REGION Network 277: SAFE OUTPUT CARD FAULT
   RUNG wire#powerrail
      Contact( "reset" )
      { S7_Templates := "SrcType := Word" } EQ_Contact(in1 := "DB101_DB_SDC_FAULTS".Carrier_Fault[28], in2 := 122)
      Coil( "DB302_HMI_Faults".Carrier28_Faults_0.%X9 )
   END_RUNG
   // the same network as SCL:
   "DB302_HMI_Faults".Carrier28_Faults_0.%X9 := "reset" AND ("DB101_DB_SDC_FAULTS".Carrier_Fault[28] = 122);
END_REGION

REGION Network 278: STANDARD INPUT CARD FAULT
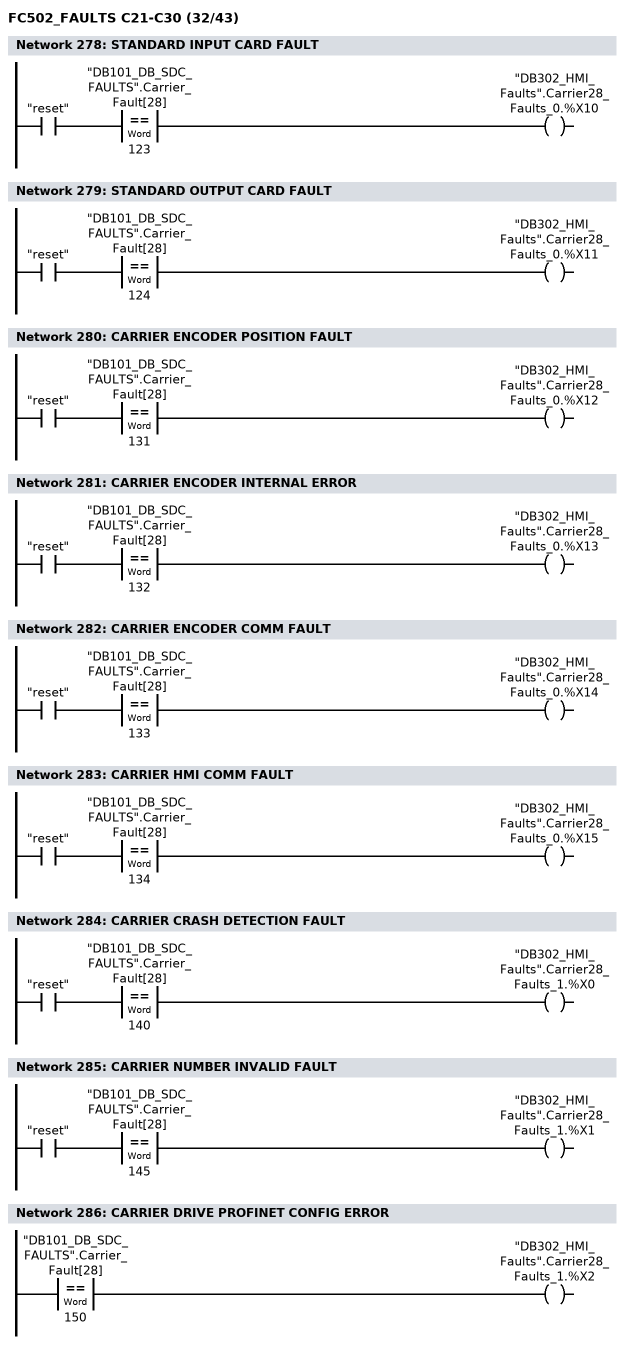
   RUNG wire#powerrail
      Contact( "reset" )
      { S7_Templates := "SrcType := Word" } EQ_Contact(in1 := "DB101_DB_SDC_FAULTS".Carrier_Fault[28], in2 := 123)
      Coil( "DB302_HMI_Faults".Carrier28_Faults_0.%X10 )
   END_RUNG
   // the same network as SCL:
   "DB302_HMI_Faults".Carrier28_Faults_0.%X10 := "reset" AND ("DB101_DB_SDC_FAULTS".Carrier_Fault[28] = 123);
END_REGION

REGION Network 279: STANDARD OUTPUT CARD FAULT
   RUNG wire#powerrail
      Contact( "reset" )
      { S7_Templates := "SrcType := Word" } EQ_Contact(in1 := "DB101_DB_SDC_FAULTS".Carrier_Fault[28], in2 := 124)
      Coil( "DB302_HMI_Faults".Carrier28_Faults_0.%X11 )
   END_RUNG
   // the same network as SCL:
   "DB302_HMI_Faults".Carrier28_Faults_0.%X11 := "reset" AND ("DB101_DB_SDC_FAULTS".Carrier_Fault[28] = 124);
END_REGION

REGION Network 280: CARRIER ENCODER POSITION FAULT
   RUNG wire#powerrail
      Contact( "reset" )
      { S7_Templates := "SrcType := Word" } EQ_Contact(in1 := "DB101_DB_SDC_FAULTS".Carrier_Fault[28], in2 := 131)
      Coil( "DB302_HMI_Faults".Carrier28_Faults_0.%X12 )
   END_RUNG
   // the same network as SCL:
   "DB302_HMI_Faults".Carrier28_Faults_0.%X12 := "reset" AND ("DB101_DB_SDC_FAULTS".Carrier_Fault[28] = 131);
END_REGION

REGION Network 281: CARRIER ENCODER INTERNAL ERROR
   RUNG wire#powerrail
      Contact( "reset" )
      { S7_Templates := "SrcType := Word" } EQ_Contact(in1 := "DB101_DB_SDC_FAULTS".Carrier_Fault[28], in2 := 132)
      Coil( "DB302_HMI_Faults".Carrier28_Faults_0.%X13 )
   END_RUNG
   // the same network as SCL:
   "DB302_HMI_Faults".Carrier28_Faults_0.%X13 := "reset" AND ("DB101_DB_SDC_FAULTS".Carrier_Fault[28] = 132);
END_REGION

REGION Network 282: CARRIER ENCODER COMM FAULT
   RUNG wire#powerrail
      Contact( "reset" )
      { S7_Templates := "SrcType := Word" } EQ_Contact(in1 := "DB101_DB_SDC_FAULTS".Carrier_Fault[28], in2 := 133)
      Coil( "DB302_HMI_Faults".Carrier28_Faults_0.%X14 )
   END_RUNG
   // the same network as SCL:
   "DB302_HMI_Faults".Carrier28_Faults_0.%X14 := "reset" AND ("DB101_DB_SDC_FAULTS".Carrier_Fault[28] = 133);
END_REGION

REGION Network 283: CARRIER HMI COMM FAULT
   RUNG wire#powerrail
      Contact( "reset" )
      { S7_Templates := "SrcType := Word" } EQ_Contact(in1 := "DB101_DB_SDC_FAULTS".Carrier_Fault[28], in2 := 134)
      Coil( "DB302_HMI_Faults".Carrier28_Faults_0.%X15 )
   END_RUNG
   // the same network as SCL:
   "DB302_HMI_Faults".Carrier28_Faults_0.%X15 := "reset" AND ("DB101_DB_SDC_FAULTS".Carrier_Fault[28] = 134);
END_REGION

REGION Network 284: CARRIER CRASH DETECTION FAULT
   RUNG wire#powerrail
      Contact( "reset" )
      { S7_Templates := "SrcType := Word" } EQ_Contact(in1 := "DB101_DB_SDC_FAULTS".Carrier_Fault[28], in2 := 140)
      Coil( "DB302_HMI_Faults".Carrier28_Faults_1.%X0 )
   END_RUNG
   // the same network as SCL:
   "DB302_HMI_Faults".Carrier28_Faults_1.%X0 := "reset" AND ("DB101_DB_SDC_FAULTS".Carrier_Fault[28] = 140);
END_REGION

REGION Network 285: CARRIER NUMBER INVALID FAULT
   RUNG wire#powerrail
      Contact( "reset" )
      { S7_Templates := "SrcType := Word" } EQ_Contact(in1 := "DB101_DB_SDC_FAULTS".Carrier_Fault[28], in2 := 145)
      Coil( "DB302_HMI_Faults".Carrier28_Faults_1.%X1 )
   END_RUNG
   // the same network as SCL:
   "DB302_HMI_Faults".Carrier28_Faults_1.%X1 := "reset" AND ("DB101_DB_SDC_FAULTS".Carrier_Fault[28] = 145);
END_REGION

REGION Network 286: CARRIER DRIVE PROFINET CONFIG ERROR
   RUNG wire#powerrail
      { S7_Templates := "SrcType := Word" } EQ_Contact(in1 := "DB101_DB_SDC_FAULTS".Carrier_Fault[28], in2 := 150)
      Coil( "DB302_HMI_Faults".Carrier28_Faults_1.%X2 )
   END_RUNG
   // the same network as SCL:
   "DB302_HMI_Faults".Carrier28_Faults_1.%X2 := "DB101_DB_SDC_FAULTS".Carrier_Fault[28] = 150;
END_REGION

REGION Network 287: CARRIER DRIVE INTERNAL COMM ERROR
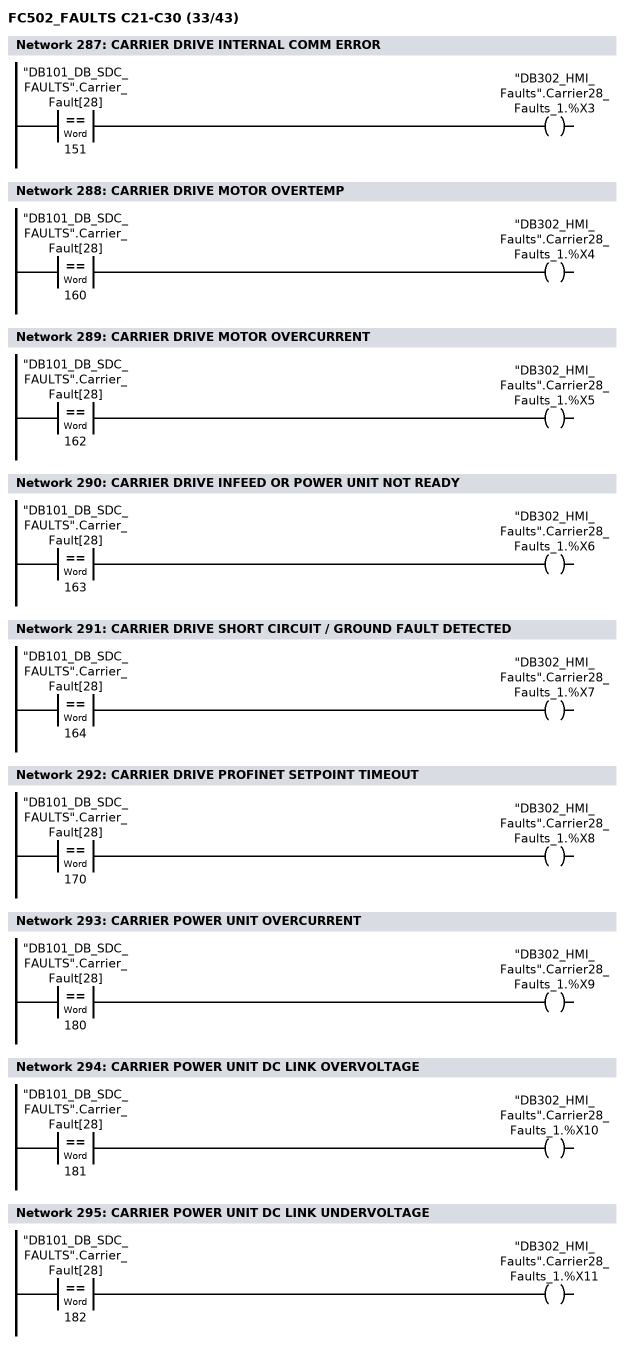
   RUNG wire#powerrail
      { S7_Templates := "SrcType := Word" } EQ_Contact(in1 := "DB101_DB_SDC_FAULTS".Carrier_Fault[28], in2 := 151)
      Coil( "DB302_HMI_Faults".Carrier28_Faults_1.%X3 )
   END_RUNG
   // the same network as SCL:
   "DB302_HMI_Faults".Carrier28_Faults_1.%X3 := "DB101_DB_SDC_FAULTS".Carrier_Fault[28] = 151;
END_REGION

REGION Network 288: CARRIER DRIVE MOTOR OVERTEMP
   RUNG wire#powerrail
      { S7_Templates := "SrcType := Word" } EQ_Contact(in1 := "DB101_DB_SDC_FAULTS".Carrier_Fault[28], in2 := 160)
      Coil( "DB302_HMI_Faults".Carrier28_Faults_1.%X4 )
   END_RUNG
   // the same network as SCL:
   "DB302_HMI_Faults".Carrier28_Faults_1.%X4 := "DB101_DB_SDC_FAULTS".Carrier_Fault[28] = 160;
END_REGION

REGION Network 289: CARRIER DRIVE MOTOR OVERCURRENT
   RUNG wire#powerrail
      { S7_Templates := "SrcType := Word" } EQ_Contact(in1 := "DB101_DB_SDC_FAULTS".Carrier_Fault[28], in2 := 162)
      Coil( "DB302_HMI_Faults".Carrier28_Faults_1.%X5 )
   END_RUNG
   // the same network as SCL:
   "DB302_HMI_Faults".Carrier28_Faults_1.%X5 := "DB101_DB_SDC_FAULTS".Carrier_Fault[28] = 162;
END_REGION

REGION Network 290: CARRIER DRIVE INFEED OR POWER UNIT NOT READY
   RUNG wire#powerrail
      { S7_Templates := "SrcType := Word" } EQ_Contact(in1 := "DB101_DB_SDC_FAULTS".Carrier_Fault[28], in2 := 163)
      Coil( "DB302_HMI_Faults".Carrier28_Faults_1.%X6 )
   END_RUNG
   // the same network as SCL:
   "DB302_HMI_Faults".Carrier28_Faults_1.%X6 := "DB101_DB_SDC_FAULTS".Carrier_Fault[28] = 163;
END_REGION

REGION Network 291: CARRIER DRIVE SHORT CIRCUIT / GROUND FAULT DETECTED
   RUNG wire#powerrail
      { S7_Templates := "SrcType := Word" } EQ_Contact(in1 := "DB101_DB_SDC_FAULTS".Carrier_Fault[28], in2 := 164)
      Coil( "DB302_HMI_Faults".Carrier28_Faults_1.%X7 )
   END_RUNG
   // the same network as SCL:
   "DB302_HMI_Faults".Carrier28_Faults_1.%X7 := "DB101_DB_SDC_FAULTS".Carrier_Fault[28] = 164;
END_REGION

REGION Network 292: CARRIER DRIVE PROFINET SETPOINT TIMEOUT
   RUNG wire#powerrail
      { S7_Templates := "SrcType := Word" } EQ_Contact(in1 := "DB101_DB_SDC_FAULTS".Carrier_Fault[28], in2 := 170)
      Coil( "DB302_HMI_Faults".Carrier28_Faults_1.%X8 )
   END_RUNG
   // the same network as SCL:
   "DB302_HMI_Faults".Carrier28_Faults_1.%X8 := "DB101_DB_SDC_FAULTS".Carrier_Fault[28] = 170;
END_REGION

REGION Network 293: CARRIER POWER UNIT OVERCURRENT
   RUNG wire#powerrail
      { S7_Templates := "SrcType := Word" } EQ_Contact(in1 := "DB101_DB_SDC_FAULTS".Carrier_Fault[28], in2 := 180)
      Coil( "DB302_HMI_Faults".Carrier28_Faults_1.%X9 )
   END_RUNG
   // the same network as SCL:
   "DB302_HMI_Faults".Carrier28_Faults_1.%X9 := "DB101_DB_SDC_FAULTS".Carrier_Fault[28] = 180;
END_REGION

REGION Network 294: CARRIER POWER UNIT DC LINK OVERVOLTAGE
   RUNG wire#powerrail
      { S7_Templates := "SrcType := Word" } EQ_Contact(in1 := "DB101_DB_SDC_FAULTS".Carrier_Fault[28], in2 := 181)
      Coil( "DB302_HMI_Faults".Carrier28_Faults_1.%X10 )
   END_RUNG
   // the same network as SCL:
   "DB302_HMI_Faults".Carrier28_Faults_1.%X10 := "DB101_DB_SDC_FAULTS".Carrier_Fault[28] = 181;
END_REGION

REGION Network 295: CARRIER POWER UNIT DC LINK UNDERVOLTAGE
   RUNG wire#powerrail
      { S7_Templates := "SrcType := Word" } EQ_Contact(in1 := "DB101_DB_SDC_FAULTS".Carrier_Fault[28], in2 := 182)
      Coil( "DB302_HMI_Faults".Carrier28_Faults_1.%X11 )
   END_RUNG
   // the same network as SCL:
   "DB302_HMI_Faults".Carrier28_Faults_1.%X11 := "DB101_DB_SDC_FAULTS".Carrier_Fault[28] = 182;
END_REGION

REGION Network 296: CARRIER POWER UNIT LINE PHASE FAILURE
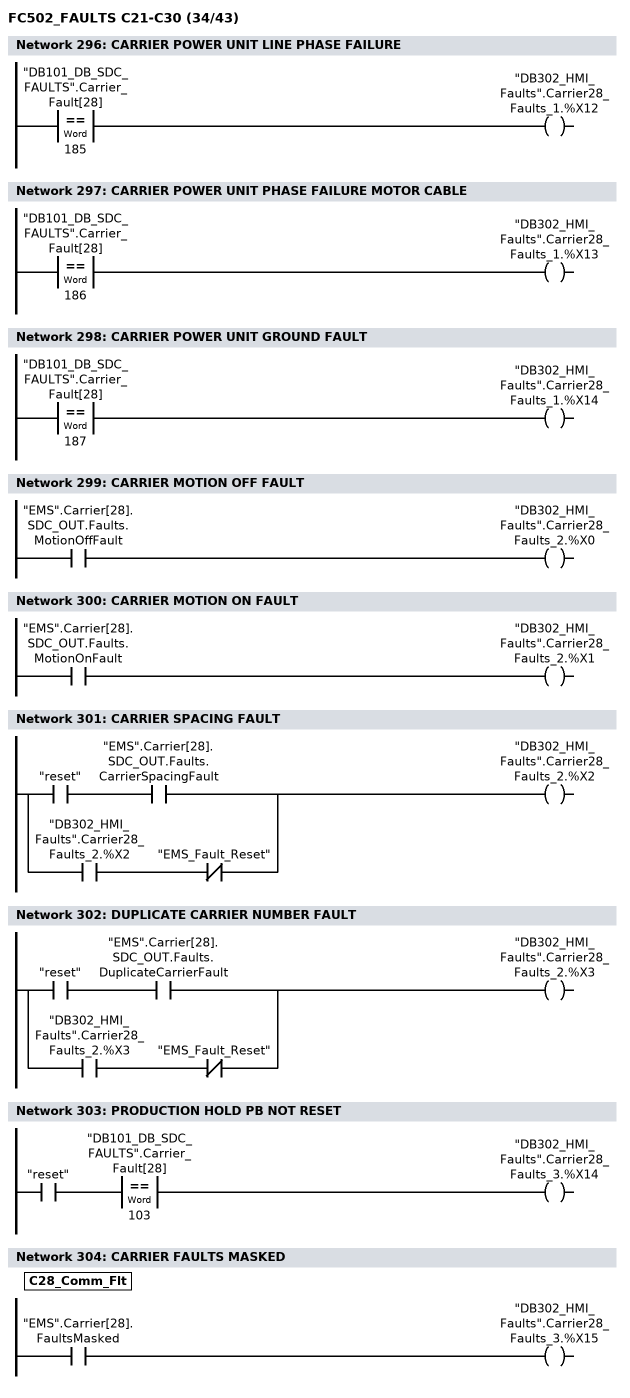
   RUNG wire#powerrail
      { S7_Templates := "SrcType := Word" } EQ_Contact(in1 := "DB101_DB_SDC_FAULTS".Carrier_Fault[28], in2 := 185)
      Coil( "DB302_HMI_Faults".Carrier28_Faults_1.%X12 )
   END_RUNG
   // the same network as SCL:
   "DB302_HMI_Faults".Carrier28_Faults_1.%X12 := "DB101_DB_SDC_FAULTS".Carrier_Fault[28] = 185;
END_REGION

REGION Network 297: CARRIER POWER UNIT PHASE FAILURE MOTOR CABLE
   RUNG wire#powerrail
      { S7_Templates := "SrcType := Word" } EQ_Contact(in1 := "DB101_DB_SDC_FAULTS".Carrier_Fault[28], in2 := 186)
      Coil( "DB302_HMI_Faults".Carrier28_Faults_1.%X13 )
   END_RUNG
   // the same network as SCL:
   "DB302_HMI_Faults".Carrier28_Faults_1.%X13 := "DB101_DB_SDC_FAULTS".Carrier_Fault[28] = 186;
END_REGION

REGION Network 298: CARRIER POWER UNIT GROUND FAULT
   RUNG wire#powerrail
      { S7_Templates := "SrcType := Word" } EQ_Contact(in1 := "DB101_DB_SDC_FAULTS".Carrier_Fault[28], in2 := 187)
      Coil( "DB302_HMI_Faults".Carrier28_Faults_1.%X14 )
   END_RUNG
   // the same network as SCL:
   "DB302_HMI_Faults".Carrier28_Faults_1.%X14 := "DB101_DB_SDC_FAULTS".Carrier_Fault[28] = 187;
END_REGION

REGION Network 299: CARRIER MOTION OFF FAULT
   RUNG wire#powerrail
      Contact( "EMS".Carrier[28].SDC_OUT.Faults.MotionOffFault )
      Coil( "DB302_HMI_Faults".Carrier28_Faults_2.%X0 )
   END_RUNG
   // the same network as SCL:
   "DB302_HMI_Faults".Carrier28_Faults_2.%X0 := "EMS".Carrier[28].SDC_OUT.Faults.MotionOffFault;
END_REGION

REGION Network 300: CARRIER MOTION ON FAULT
   RUNG wire#powerrail
      Contact( "EMS".Carrier[28].SDC_OUT.Faults.MotionOnFault )
      Coil( "DB302_HMI_Faults".Carrier28_Faults_2.%X1 )
   END_RUNG
   // the same network as SCL:
   "DB302_HMI_Faults".Carrier28_Faults_2.%X1 := "EMS".Carrier[28].SDC_OUT.Faults.MotionOnFault;
END_REGION

REGION Network 301: CARRIER SPACING FAULT
   RUNG wire#powerrail
      Contact( "reset" )
      Contact( "EMS".Carrier[28].SDC_OUT.Faults.CarrierSpacingFault )
      wire#w1
      Coil( "DB302_HMI_Faults".Carrier28_Faults_2.%X2 )
   END_RUNG
   RUNG wire#powerrail
      Contact( "DB302_HMI_Faults".Carrier28_Faults_2.%X2 )
      I_Contact( "EMS_Fault_Reset" )
   END_RUNG wire#w1
   // the same network as SCL:
   "DB302_HMI_Faults".Carrier28_Faults_2.%X2 := ("reset" AND "EMS".Carrier[28].SDC_OUT.Faults.CarrierSpacingFault) OR ("DB302_HMI_Faults".Carrier28_Faults_2.%X2 AND NOT "EMS_Fault_Reset");
END_REGION

REGION Network 302: DUPLICATE CARRIER NUMBER FAULT
   RUNG wire#powerrail
      Contact( "reset" )
      Contact( "EMS".Carrier[28].SDC_OUT.Faults.DuplicateCarrierFault )
      wire#w1
      Coil( "DB302_HMI_Faults".Carrier28_Faults_2.%X3 )
   END_RUNG
   RUNG wire#powerrail
      Contact( "DB302_HMI_Faults".Carrier28_Faults_2.%X3 )
      I_Contact( "EMS_Fault_Reset" )
   END_RUNG wire#w1
   // the same network as SCL:
   "DB302_HMI_Faults".Carrier28_Faults_2.%X3 := ("reset" AND "EMS".Carrier[28].SDC_OUT.Faults.DuplicateCarrierFault) OR ("DB302_HMI_Faults".Carrier28_Faults_2.%X3 AND NOT "EMS_Fault_Reset");
END_REGION

REGION Network 303: PRODUCTION HOLD PB NOT RESET
   RUNG wire#powerrail
      Contact( "reset" )
      { S7_Templates := "SrcType := Word" } EQ_Contact(in1 := "DB101_DB_SDC_FAULTS".Carrier_Fault[28], in2 := 103)
      Coil( "DB302_HMI_Faults".Carrier28_Faults_3.%X14 )
   END_RUNG
   // the same network as SCL:
   "DB302_HMI_Faults".Carrier28_Faults_3.%X14 := "reset" AND ("DB101_DB_SDC_FAULTS".Carrier_Fault[28] = 103);
END_REGION

REGION Network 304: CARRIER FAULTS MASKED
   Label( C28_Comm_Flt )
   RUNG wire#powerrail
      Contact( "EMS".Carrier[28].FaultsMasked )
      Coil( "DB302_HMI_Faults".Carrier28_Faults_3.%X15 )
   END_RUNG
   // the same network as SCL:
   C28_Comm_Flt:
   "DB302_HMI_Faults".Carrier28_Faults_3.%X15 := "EMS".Carrier[28].FaultsMasked;
END_REGION

REGION Network 305: CARRIER 29 FAULTS
END_REGION

REGION Network 306: CARRIER PLC NOT COMMUNICATING
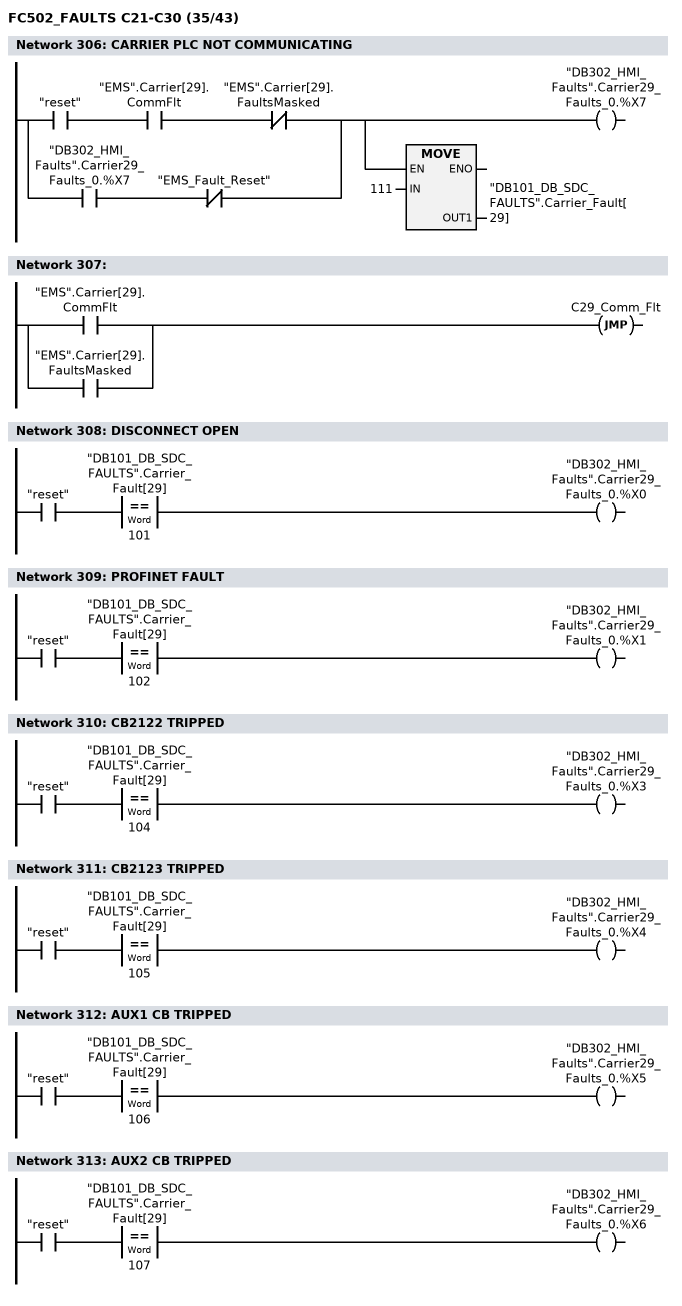
   RUNG wire#powerrail
      Contact( "reset" )
      Contact( "EMS".Carrier[29].CommFlt )
      I_Contact( "EMS".Carrier[29].FaultsMasked )
      wire#w1
      Coil( "DB302_HMI_Faults".Carrier29_Faults_0.%X7 )
   END_RUNG
   RUNG wire#powerrail
      Contact( "DB302_HMI_Faults".Carrier29_Faults_0.%X7 )
      I_Contact( "EMS_Fault_Reset" )
   END_RUNG wire#w1
   RUNG wire#w1
      Move(in := 111, out1 => "DB101_DB_SDC_FAULTS".Carrier_Fault[29])
   END_RUNG
   // the same network as SCL:
   "DB302_HMI_Faults".Carrier29_Faults_0.%X7 := ("reset" AND "EMS".Carrier[29].CommFlt AND NOT "EMS".Carrier[29].FaultsMasked) OR ("DB302_HMI_Faults".Carrier29_Faults_0.%X7 AND NOT "EMS_Fault_Reset");
   IF "DB302_HMI_Faults".Carrier29_Faults_0.%X7 THEN "DB101_DB_SDC_FAULTS".Carrier_Fault[29] := 111; END_IF;
END_REGION

REGION Network 307
   RUNG wire#powerrail
      Contact( "EMS".Carrier[29].CommFlt )
      wire#w1
      JumpCoil( C29_Comm_Flt )
   END_RUNG
   RUNG wire#powerrail
      Contact( "EMS".Carrier[29].FaultsMasked )
   END_RUNG wire#w1
   // the same network as SCL:
   IF "EMS".Carrier[29].CommFlt OR "EMS".Carrier[29].FaultsMasked THEN GOTO C29_Comm_Flt; END_IF;
END_REGION

REGION Network 308: DISCONNECT OPEN
   RUNG wire#powerrail
      Contact( "reset" )
      { S7_Templates := "SrcType := Word" } EQ_Contact(in1 := "DB101_DB_SDC_FAULTS".Carrier_Fault[29], in2 := 101)
      Coil( "DB302_HMI_Faults".Carrier29_Faults_0.%X0 )
   END_RUNG
   // the same network as SCL:
   "DB302_HMI_Faults".Carrier29_Faults_0.%X0 := "reset" AND ("DB101_DB_SDC_FAULTS".Carrier_Fault[29] = 101);
END_REGION

REGION Network 309: PROFINET FAULT
   RUNG wire#powerrail
      Contact( "reset" )
      { S7_Templates := "SrcType := Word" } EQ_Contact(in1 := "DB101_DB_SDC_FAULTS".Carrier_Fault[29], in2 := 102)
      Coil( "DB302_HMI_Faults".Carrier29_Faults_0.%X1 )
   END_RUNG
   // the same network as SCL:
   "DB302_HMI_Faults".Carrier29_Faults_0.%X1 := "reset" AND ("DB101_DB_SDC_FAULTS".Carrier_Fault[29] = 102);
END_REGION

REGION Network 310: CB2122 TRIPPED
   RUNG wire#powerrail
      Contact( "reset" )
      { S7_Templates := "SrcType := Word" } EQ_Contact(in1 := "DB101_DB_SDC_FAULTS".Carrier_Fault[29], in2 := 104)
      Coil( "DB302_HMI_Faults".Carrier29_Faults_0.%X3 )
   END_RUNG
   // the same network as SCL:
   "DB302_HMI_Faults".Carrier29_Faults_0.%X3 := "reset" AND ("DB101_DB_SDC_FAULTS".Carrier_Fault[29] = 104);
END_REGION

REGION Network 311: CB2123 TRIPPED
   RUNG wire#powerrail
      Contact( "reset" )
      { S7_Templates := "SrcType := Word" } EQ_Contact(in1 := "DB101_DB_SDC_FAULTS".Carrier_Fault[29], in2 := 105)
      Coil( "DB302_HMI_Faults".Carrier29_Faults_0.%X4 )
   END_RUNG
   // the same network as SCL:
   "DB302_HMI_Faults".Carrier29_Faults_0.%X4 := "reset" AND ("DB101_DB_SDC_FAULTS".Carrier_Fault[29] = 105);
END_REGION

REGION Network 312: AUX1 CB TRIPPED
   RUNG wire#powerrail
      Contact( "reset" )
      { S7_Templates := "SrcType := Word" } EQ_Contact(in1 := "DB101_DB_SDC_FAULTS".Carrier_Fault[29], in2 := 106)
      Coil( "DB302_HMI_Faults".Carrier29_Faults_0.%X5 )
   END_RUNG
   // the same network as SCL:
   "DB302_HMI_Faults".Carrier29_Faults_0.%X5 := "reset" AND ("DB101_DB_SDC_FAULTS".Carrier_Fault[29] = 106);
END_REGION

REGION Network 313: AUX2 CB TRIPPED
   RUNG wire#powerrail
      Contact( "reset" )
      { S7_Templates := "SrcType := Word" } EQ_Contact(in1 := "DB101_DB_SDC_FAULTS".Carrier_Fault[29], in2 := 107)
      Coil( "DB302_HMI_Faults".Carrier29_Faults_0.%X6 )
   END_RUNG
   // the same network as SCL:
   "DB302_HMI_Faults".Carrier29_Faults_0.%X6 := "reset" AND ("DB101_DB_SDC_FAULTS".Carrier_Fault[29] = 107);
END_REGION

REGION Network 314: SAFE INPUT CARD FAULT
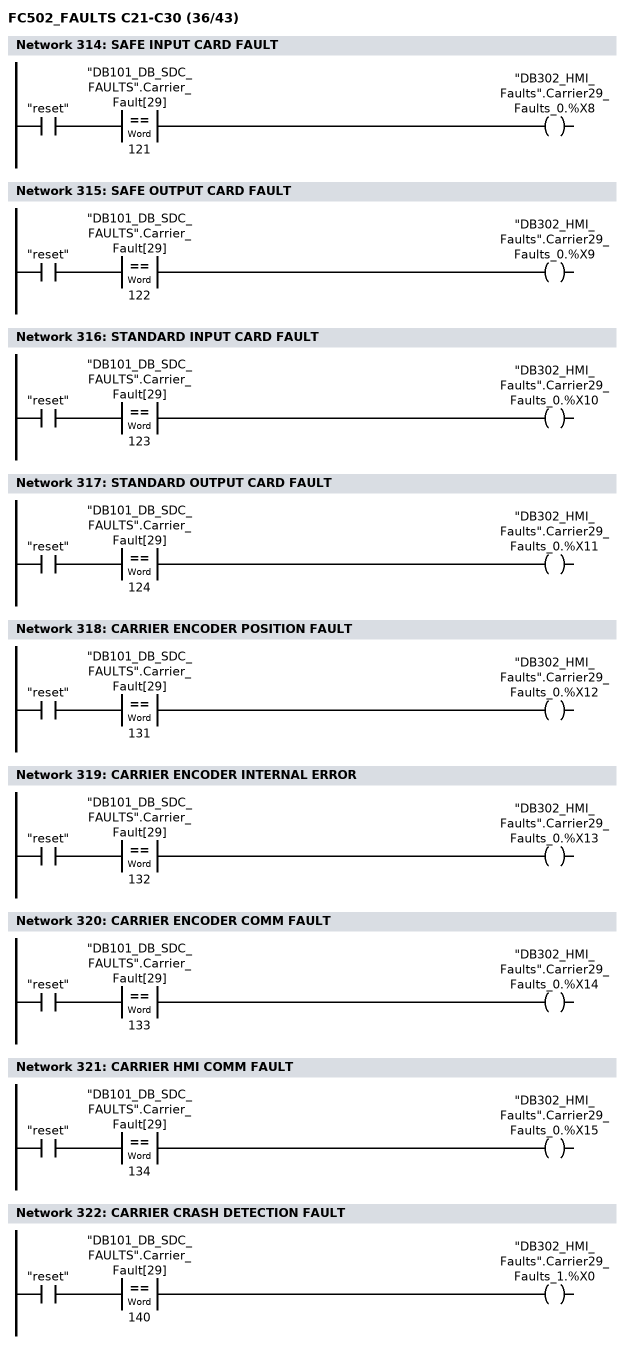
   RUNG wire#powerrail
      Contact( "reset" )
      { S7_Templates := "SrcType := Word" } EQ_Contact(in1 := "DB101_DB_SDC_FAULTS".Carrier_Fault[29], in2 := 121)
      Coil( "DB302_HMI_Faults".Carrier29_Faults_0.%X8 )
   END_RUNG
   // the same network as SCL:
   "DB302_HMI_Faults".Carrier29_Faults_0.%X8 := "reset" AND ("DB101_DB_SDC_FAULTS".Carrier_Fault[29] = 121);
END_REGION

REGION Network 315: SAFE OUTPUT CARD FAULT
   RUNG wire#powerrail
      Contact( "reset" )
      { S7_Templates := "SrcType := Word" } EQ_Contact(in1 := "DB101_DB_SDC_FAULTS".Carrier_Fault[29], in2 := 122)
      Coil( "DB302_HMI_Faults".Carrier29_Faults_0.%X9 )
   END_RUNG
   // the same network as SCL:
   "DB302_HMI_Faults".Carrier29_Faults_0.%X9 := "reset" AND ("DB101_DB_SDC_FAULTS".Carrier_Fault[29] = 122);
END_REGION

REGION Network 316: STANDARD INPUT CARD FAULT
   RUNG wire#powerrail
      Contact( "reset" )
      { S7_Templates := "SrcType := Word" } EQ_Contact(in1 := "DB101_DB_SDC_FAULTS".Carrier_Fault[29], in2 := 123)
      Coil( "DB302_HMI_Faults".Carrier29_Faults_0.%X10 )
   END_RUNG
   // the same network as SCL:
   "DB302_HMI_Faults".Carrier29_Faults_0.%X10 := "reset" AND ("DB101_DB_SDC_FAULTS".Carrier_Fault[29] = 123);
END_REGION

REGION Network 317: STANDARD OUTPUT CARD FAULT
   RUNG wire#powerrail
      Contact( "reset" )
      { S7_Templates := "SrcType := Word" } EQ_Contact(in1 := "DB101_DB_SDC_FAULTS".Carrier_Fault[29], in2 := 124)
      Coil( "DB302_HMI_Faults".Carrier29_Faults_0.%X11 )
   END_RUNG
   // the same network as SCL:
   "DB302_HMI_Faults".Carrier29_Faults_0.%X11 := "reset" AND ("DB101_DB_SDC_FAULTS".Carrier_Fault[29] = 124);
END_REGION

REGION Network 318: CARRIER ENCODER POSITION FAULT
   RUNG wire#powerrail
      Contact( "reset" )
      { S7_Templates := "SrcType := Word" } EQ_Contact(in1 := "DB101_DB_SDC_FAULTS".Carrier_Fault[29], in2 := 131)
      Coil( "DB302_HMI_Faults".Carrier29_Faults_0.%X12 )
   END_RUNG
   // the same network as SCL:
   "DB302_HMI_Faults".Carrier29_Faults_0.%X12 := "reset" AND ("DB101_DB_SDC_FAULTS".Carrier_Fault[29] = 131);
END_REGION

REGION Network 319: CARRIER ENCODER INTERNAL ERROR
   RUNG wire#powerrail
      Contact( "reset" )
      { S7_Templates := "SrcType := Word" } EQ_Contact(in1 := "DB101_DB_SDC_FAULTS".Carrier_Fault[29], in2 := 132)
      Coil( "DB302_HMI_Faults".Carrier29_Faults_0.%X13 )
   END_RUNG
   // the same network as SCL:
   "DB302_HMI_Faults".Carrier29_Faults_0.%X13 := "reset" AND ("DB101_DB_SDC_FAULTS".Carrier_Fault[29] = 132);
END_REGION

REGION Network 320: CARRIER ENCODER COMM FAULT
   RUNG wire#powerrail
      Contact( "reset" )
      { S7_Templates := "SrcType := Word" } EQ_Contact(in1 := "DB101_DB_SDC_FAULTS".Carrier_Fault[29], in2 := 133)
      Coil( "DB302_HMI_Faults".Carrier29_Faults_0.%X14 )
   END_RUNG
   // the same network as SCL:
   "DB302_HMI_Faults".Carrier29_Faults_0.%X14 := "reset" AND ("DB101_DB_SDC_FAULTS".Carrier_Fault[29] = 133);
END_REGION

REGION Network 321: CARRIER HMI COMM FAULT
   RUNG wire#powerrail
      Contact( "reset" )
      { S7_Templates := "SrcType := Word" } EQ_Contact(in1 := "DB101_DB_SDC_FAULTS".Carrier_Fault[29], in2 := 134)
      Coil( "DB302_HMI_Faults".Carrier29_Faults_0.%X15 )
   END_RUNG
   // the same network as SCL:
   "DB302_HMI_Faults".Carrier29_Faults_0.%X15 := "reset" AND ("DB101_DB_SDC_FAULTS".Carrier_Fault[29] = 134);
END_REGION

REGION Network 322: CARRIER CRASH DETECTION FAULT
   RUNG wire#powerrail
      Contact( "reset" )
      { S7_Templates := "SrcType := Word" } EQ_Contact(in1 := "DB101_DB_SDC_FAULTS".Carrier_Fault[29], in2 := 140)
      Coil( "DB302_HMI_Faults".Carrier29_Faults_1.%X0 )
   END_RUNG
   // the same network as SCL:
   "DB302_HMI_Faults".Carrier29_Faults_1.%X0 := "reset" AND ("DB101_DB_SDC_FAULTS".Carrier_Fault[29] = 140);
END_REGION

REGION Network 323: CARRIER NUMBER INVALID FAULT
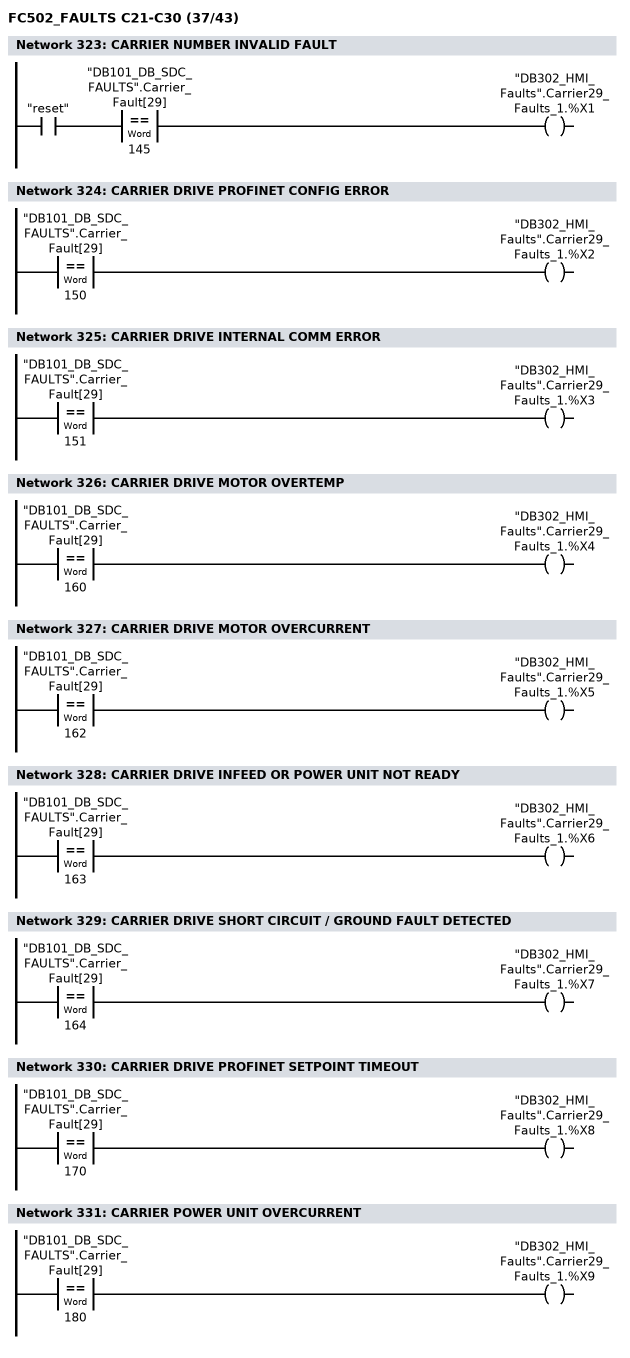
   RUNG wire#powerrail
      Contact( "reset" )
      { S7_Templates := "SrcType := Word" } EQ_Contact(in1 := "DB101_DB_SDC_FAULTS".Carrier_Fault[29], in2 := 145)
      Coil( "DB302_HMI_Faults".Carrier29_Faults_1.%X1 )
   END_RUNG
   // the same network as SCL:
   "DB302_HMI_Faults".Carrier29_Faults_1.%X1 := "reset" AND ("DB101_DB_SDC_FAULTS".Carrier_Fault[29] = 145);
END_REGION

REGION Network 324: CARRIER DRIVE PROFINET CONFIG ERROR
   RUNG wire#powerrail
      { S7_Templates := "SrcType := Word" } EQ_Contact(in1 := "DB101_DB_SDC_FAULTS".Carrier_Fault[29], in2 := 150)
      Coil( "DB302_HMI_Faults".Carrier29_Faults_1.%X2 )
   END_RUNG
   // the same network as SCL:
   "DB302_HMI_Faults".Carrier29_Faults_1.%X2 := "DB101_DB_SDC_FAULTS".Carrier_Fault[29] = 150;
END_REGION

REGION Network 325: CARRIER DRIVE INTERNAL COMM ERROR
   RUNG wire#powerrail
      { S7_Templates := "SrcType := Word" } EQ_Contact(in1 := "DB101_DB_SDC_FAULTS".Carrier_Fault[29], in2 := 151)
      Coil( "DB302_HMI_Faults".Carrier29_Faults_1.%X3 )
   END_RUNG
   // the same network as SCL:
   "DB302_HMI_Faults".Carrier29_Faults_1.%X3 := "DB101_DB_SDC_FAULTS".Carrier_Fault[29] = 151;
END_REGION

REGION Network 326: CARRIER DRIVE MOTOR OVERTEMP
   RUNG wire#powerrail
      { S7_Templates := "SrcType := Word" } EQ_Contact(in1 := "DB101_DB_SDC_FAULTS".Carrier_Fault[29], in2 := 160)
      Coil( "DB302_HMI_Faults".Carrier29_Faults_1.%X4 )
   END_RUNG
   // the same network as SCL:
   "DB302_HMI_Faults".Carrier29_Faults_1.%X4 := "DB101_DB_SDC_FAULTS".Carrier_Fault[29] = 160;
END_REGION

REGION Network 327: CARRIER DRIVE MOTOR OVERCURRENT
   RUNG wire#powerrail
      { S7_Templates := "SrcType := Word" } EQ_Contact(in1 := "DB101_DB_SDC_FAULTS".Carrier_Fault[29], in2 := 162)
      Coil( "DB302_HMI_Faults".Carrier29_Faults_1.%X5 )
   END_RUNG
   // the same network as SCL:
   "DB302_HMI_Faults".Carrier29_Faults_1.%X5 := "DB101_DB_SDC_FAULTS".Carrier_Fault[29] = 162;
END_REGION

REGION Network 328: CARRIER DRIVE INFEED OR POWER UNIT NOT READY
   RUNG wire#powerrail
      { S7_Templates := "SrcType := Word" } EQ_Contact(in1 := "DB101_DB_SDC_FAULTS".Carrier_Fault[29], in2 := 163)
      Coil( "DB302_HMI_Faults".Carrier29_Faults_1.%X6 )
   END_RUNG
   // the same network as SCL:
   "DB302_HMI_Faults".Carrier29_Faults_1.%X6 := "DB101_DB_SDC_FAULTS".Carrier_Fault[29] = 163;
END_REGION

REGION Network 329: CARRIER DRIVE SHORT CIRCUIT / GROUND FAULT DETECTED
   RUNG wire#powerrail
      { S7_Templates := "SrcType := Word" } EQ_Contact(in1 := "DB101_DB_SDC_FAULTS".Carrier_Fault[29], in2 := 164)
      Coil( "DB302_HMI_Faults".Carrier29_Faults_1.%X7 )
   END_RUNG
   // the same network as SCL:
   "DB302_HMI_Faults".Carrier29_Faults_1.%X7 := "DB101_DB_SDC_FAULTS".Carrier_Fault[29] = 164;
END_REGION

REGION Network 330: CARRIER DRIVE PROFINET SETPOINT TIMEOUT
   RUNG wire#powerrail
      { S7_Templates := "SrcType := Word" } EQ_Contact(in1 := "DB101_DB_SDC_FAULTS".Carrier_Fault[29], in2 := 170)
      Coil( "DB302_HMI_Faults".Carrier29_Faults_1.%X8 )
   END_RUNG
   // the same network as SCL:
   "DB302_HMI_Faults".Carrier29_Faults_1.%X8 := "DB101_DB_SDC_FAULTS".Carrier_Fault[29] = 170;
END_REGION

REGION Network 331: CARRIER POWER UNIT OVERCURRENT
   RUNG wire#powerrail
      { S7_Templates := "SrcType := Word" } EQ_Contact(in1 := "DB101_DB_SDC_FAULTS".Carrier_Fault[29], in2 := 180)
      Coil( "DB302_HMI_Faults".Carrier29_Faults_1.%X9 )
   END_RUNG
   // the same network as SCL:
   "DB302_HMI_Faults".Carrier29_Faults_1.%X9 := "DB101_DB_SDC_FAULTS".Carrier_Fault[29] = 180;
END_REGION

REGION Network 332: CARRIER POWER UNIT DC LINK OVERVOLTAGE
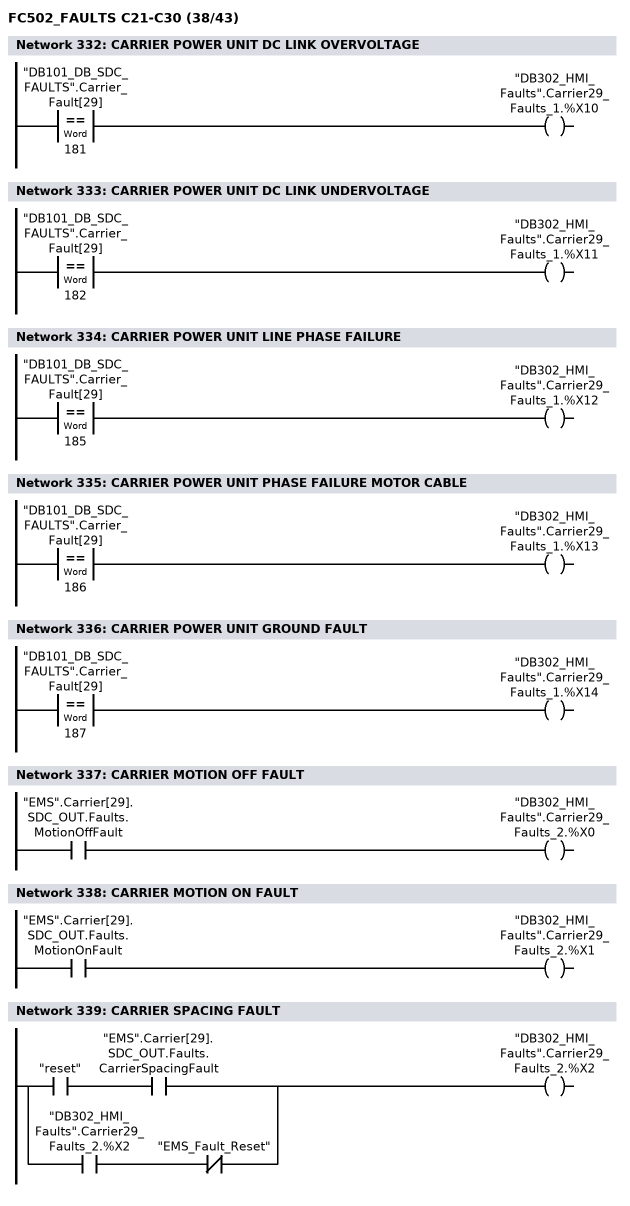
   RUNG wire#powerrail
      { S7_Templates := "SrcType := Word" } EQ_Contact(in1 := "DB101_DB_SDC_FAULTS".Carrier_Fault[29], in2 := 181)
      Coil( "DB302_HMI_Faults".Carrier29_Faults_1.%X10 )
   END_RUNG
   // the same network as SCL:
   "DB302_HMI_Faults".Carrier29_Faults_1.%X10 := "DB101_DB_SDC_FAULTS".Carrier_Fault[29] = 181;
END_REGION

REGION Network 333: CARRIER POWER UNIT DC LINK UNDERVOLTAGE
   RUNG wire#powerrail
      { S7_Templates := "SrcType := Word" } EQ_Contact(in1 := "DB101_DB_SDC_FAULTS".Carrier_Fault[29], in2 := 182)
      Coil( "DB302_HMI_Faults".Carrier29_Faults_1.%X11 )
   END_RUNG
   // the same network as SCL:
   "DB302_HMI_Faults".Carrier29_Faults_1.%X11 := "DB101_DB_SDC_FAULTS".Carrier_Fault[29] = 182;
END_REGION

REGION Network 334: CARRIER POWER UNIT LINE PHASE FAILURE
   RUNG wire#powerrail
      { S7_Templates := "SrcType := Word" } EQ_Contact(in1 := "DB101_DB_SDC_FAULTS".Carrier_Fault[29], in2 := 185)
      Coil( "DB302_HMI_Faults".Carrier29_Faults_1.%X12 )
   END_RUNG
   // the same network as SCL:
   "DB302_HMI_Faults".Carrier29_Faults_1.%X12 := "DB101_DB_SDC_FAULTS".Carrier_Fault[29] = 185;
END_REGION

REGION Network 335: CARRIER POWER UNIT PHASE FAILURE MOTOR CABLE
   RUNG wire#powerrail
      { S7_Templates := "SrcType := Word" } EQ_Contact(in1 := "DB101_DB_SDC_FAULTS".Carrier_Fault[29], in2 := 186)
      Coil( "DB302_HMI_Faults".Carrier29_Faults_1.%X13 )
   END_RUNG
   // the same network as SCL:
   "DB302_HMI_Faults".Carrier29_Faults_1.%X13 := "DB101_DB_SDC_FAULTS".Carrier_Fault[29] = 186;
END_REGION

REGION Network 336: CARRIER POWER UNIT GROUND FAULT
   RUNG wire#powerrail
      { S7_Templates := "SrcType := Word" } EQ_Contact(in1 := "DB101_DB_SDC_FAULTS".Carrier_Fault[29], in2 := 187)
      Coil( "DB302_HMI_Faults".Carrier29_Faults_1.%X14 )
   END_RUNG
   // the same network as SCL:
   "DB302_HMI_Faults".Carrier29_Faults_1.%X14 := "DB101_DB_SDC_FAULTS".Carrier_Fault[29] = 187;
END_REGION

REGION Network 337: CARRIER MOTION OFF FAULT
   RUNG wire#powerrail
      Contact( "EMS".Carrier[29].SDC_OUT.Faults.MotionOffFault )
      Coil( "DB302_HMI_Faults".Carrier29_Faults_2.%X0 )
   END_RUNG
   // the same network as SCL:
   "DB302_HMI_Faults".Carrier29_Faults_2.%X0 := "EMS".Carrier[29].SDC_OUT.Faults.MotionOffFault;
END_REGION

REGION Network 338: CARRIER MOTION ON FAULT
   RUNG wire#powerrail
      Contact( "EMS".Carrier[29].SDC_OUT.Faults.MotionOnFault )
      Coil( "DB302_HMI_Faults".Carrier29_Faults_2.%X1 )
   END_RUNG
   // the same network as SCL:
   "DB302_HMI_Faults".Carrier29_Faults_2.%X1 := "EMS".Carrier[29].SDC_OUT.Faults.MotionOnFault;
END_REGION

REGION Network 339: CARRIER SPACING FAULT
   RUNG wire#powerrail
      Contact( "reset" )
      Contact( "EMS".Carrier[29].SDC_OUT.Faults.CarrierSpacingFault )
      wire#w1
      Coil( "DB302_HMI_Faults".Carrier29_Faults_2.%X2 )
   END_RUNG
   RUNG wire#powerrail
      Contact( "DB302_HMI_Faults".Carrier29_Faults_2.%X2 )
      I_Contact( "EMS_Fault_Reset" )
   END_RUNG wire#w1
   // the same network as SCL:
   "DB302_HMI_Faults".Carrier29_Faults_2.%X2 := ("reset" AND "EMS".Carrier[29].SDC_OUT.Faults.CarrierSpacingFault) OR ("DB302_HMI_Faults".Carrier29_Faults_2.%X2 AND NOT "EMS_Fault_Reset");
END_REGION

REGION Network 340: DUPLICATE CARRIER NUMBER FAULT
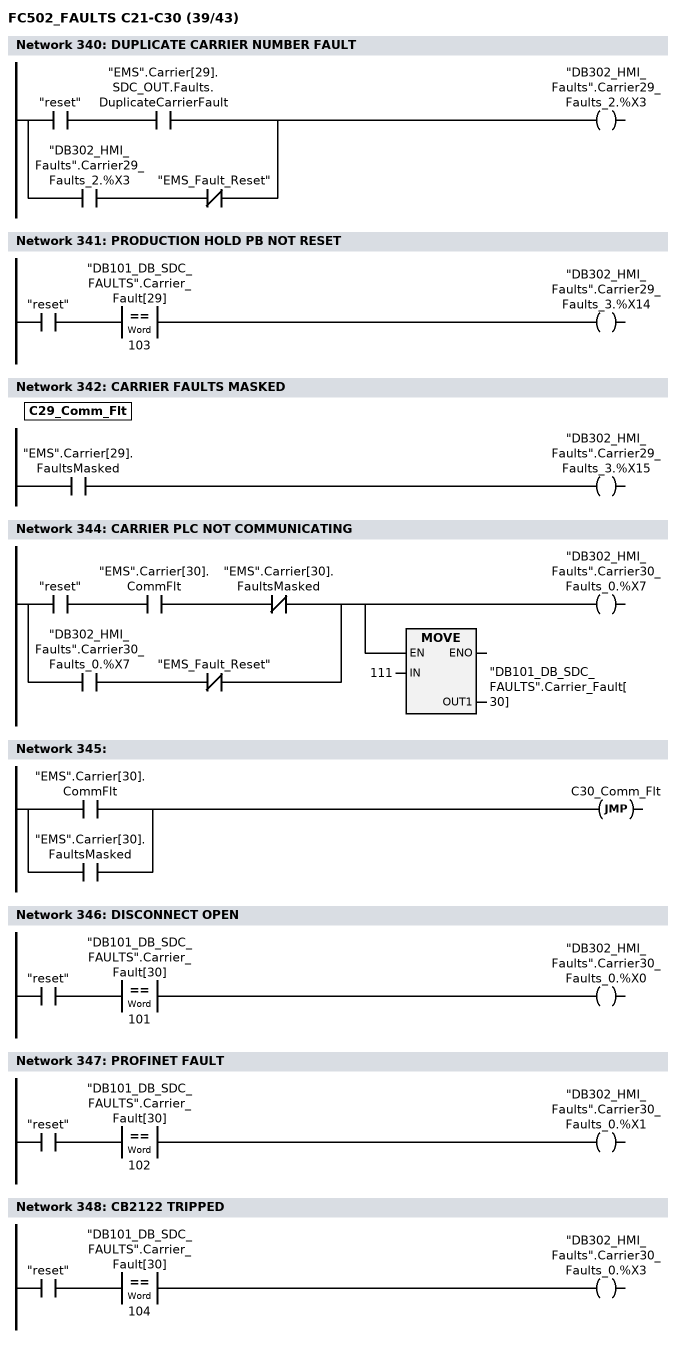
   RUNG wire#powerrail
      Contact( "reset" )
      Contact( "EMS".Carrier[29].SDC_OUT.Faults.DuplicateCarrierFault )
      wire#w1
      Coil( "DB302_HMI_Faults".Carrier29_Faults_2.%X3 )
   END_RUNG
   RUNG wire#powerrail
      Contact( "DB302_HMI_Faults".Carrier29_Faults_2.%X3 )
      I_Contact( "EMS_Fault_Reset" )
   END_RUNG wire#w1
   // the same network as SCL:
   "DB302_HMI_Faults".Carrier29_Faults_2.%X3 := ("reset" AND "EMS".Carrier[29].SDC_OUT.Faults.DuplicateCarrierFault) OR ("DB302_HMI_Faults".Carrier29_Faults_2.%X3 AND NOT "EMS_Fault_Reset");
END_REGION

REGION Network 341: PRODUCTION HOLD PB NOT RESET
   RUNG wire#powerrail
      Contact( "reset" )
      { S7_Templates := "SrcType := Word" } EQ_Contact(in1 := "DB101_DB_SDC_FAULTS".Carrier_Fault[29], in2 := 103)
      Coil( "DB302_HMI_Faults".Carrier29_Faults_3.%X14 )
   END_RUNG
   // the same network as SCL:
   "DB302_HMI_Faults".Carrier29_Faults_3.%X14 := "reset" AND ("DB101_DB_SDC_FAULTS".Carrier_Fault[29] = 103);
END_REGION

REGION Network 342: CARRIER FAULTS MASKED
   Label( C29_Comm_Flt )
   RUNG wire#powerrail
      Contact( "EMS".Carrier[29].FaultsMasked )
      Coil( "DB302_HMI_Faults".Carrier29_Faults_3.%X15 )
   END_RUNG
   // the same network as SCL:
   C29_Comm_Flt:
   "DB302_HMI_Faults".Carrier29_Faults_3.%X15 := "EMS".Carrier[29].FaultsMasked;
END_REGION

REGION Network 343: CARRIER 30 FAULTS
END_REGION

REGION Network 344: CARRIER PLC NOT COMMUNICATING
   RUNG wire#powerrail
      Contact( "reset" )
      Contact( "EMS".Carrier[30].CommFlt )
      I_Contact( "EMS".Carrier[30].FaultsMasked )
      wire#w1
      Coil( "DB302_HMI_Faults".Carrier30_Faults_0.%X7 )
   END_RUNG
   RUNG wire#powerrail
      Contact( "DB302_HMI_Faults".Carrier30_Faults_0.%X7 )
      I_Contact( "EMS_Fault_Reset" )
   END_RUNG wire#w1
   RUNG wire#w1
      Move(in := 111, out1 => "DB101_DB_SDC_FAULTS".Carrier_Fault[30])
   END_RUNG
   // the same network as SCL:
   "DB302_HMI_Faults".Carrier30_Faults_0.%X7 := ("reset" AND "EMS".Carrier[30].CommFlt AND NOT "EMS".Carrier[30].FaultsMasked) OR ("DB302_HMI_Faults".Carrier30_Faults_0.%X7 AND NOT "EMS_Fault_Reset");
   IF "DB302_HMI_Faults".Carrier30_Faults_0.%X7 THEN "DB101_DB_SDC_FAULTS".Carrier_Fault[30] := 111; END_IF;
END_REGION

REGION Network 345
   RUNG wire#powerrail
      Contact( "EMS".Carrier[30].CommFlt )
      wire#w1
      JumpCoil( C30_Comm_Flt )
   END_RUNG
   RUNG wire#powerrail
      Contact( "EMS".Carrier[30].FaultsMasked )
   END_RUNG wire#w1
   // the same network as SCL:
   IF "EMS".Carrier[30].CommFlt OR "EMS".Carrier[30].FaultsMasked THEN GOTO C30_Comm_Flt; END_IF;
END_REGION

REGION Network 346: DISCONNECT OPEN
   RUNG wire#powerrail
      Contact( "reset" )
      { S7_Templates := "SrcType := Word" } EQ_Contact(in1 := "DB101_DB_SDC_FAULTS".Carrier_Fault[30], in2 := 101)
      Coil( "DB302_HMI_Faults".Carrier30_Faults_0.%X0 )
   END_RUNG
   // the same network as SCL:
   "DB302_HMI_Faults".Carrier30_Faults_0.%X0 := "reset" AND ("DB101_DB_SDC_FAULTS".Carrier_Fault[30] = 101);
END_REGION

REGION Network 347: PROFINET FAULT
   RUNG wire#powerrail
      Contact( "reset" )
      { S7_Templates := "SrcType := Word" } EQ_Contact(in1 := "DB101_DB_SDC_FAULTS".Carrier_Fault[30], in2 := 102)
      Coil( "DB302_HMI_Faults".Carrier30_Faults_0.%X1 )
   END_RUNG
   // the same network as SCL:
   "DB302_HMI_Faults".Carrier30_Faults_0.%X1 := "reset" AND ("DB101_DB_SDC_FAULTS".Carrier_Fault[30] = 102);
END_REGION

REGION Network 348: CB2122 TRIPPED
   RUNG wire#powerrail
      Contact( "reset" )
      { S7_Templates := "SrcType := Word" } EQ_Contact(in1 := "DB101_DB_SDC_FAULTS".Carrier_Fault[30], in2 := 104)
      Coil( "DB302_HMI_Faults".Carrier30_Faults_0.%X3 )
   END_RUNG
   // the same network as SCL:
   "DB302_HMI_Faults".Carrier30_Faults_0.%X3 := "reset" AND ("DB101_DB_SDC_FAULTS".Carrier_Fault[30] = 104);
END_REGION

REGION Network 349: CB2123 TRIPPED
